// TIA Portal project "EbAndon v2_1_0" (V15) (continued)
   // me.stations[14] : chm 04
   // me.stations[15] : cdo 01
   // me.stations[16] : cdo 02
   // me.stations[17] : cdo 03
   // me.stations[18] : bfl 01
   // me.stations[19] : bfl 02
   // me.stations[20] : bfl 03
   // me.stations[21] : lgs 01
   // me.stations[22] : lgs 02
   // me.stations[23] : lgs 03
   // me.stations[24] : cv 01
   // me.stations[25] : cv 02
   // me.stations[26] : cv 03
   // me.stations[27] : cv 04
   // me.stations[28] : pc 01
   // me.stations[29] : pc 02
END_DATA_BLOCK

// folder: Network Diagnostics

DATA_BLOCK "Net Diag: Global"   // DB7
{ S7_Optimized_Access := 'TRUE' }
VERSION : 0.1
   VAR
      plcData : "UserDiag_typePLC";   // PLC diagnostics data
      ioSystemData : Array[1.."USERDIAG_IO_SYSTEMS_UPPER_LIM"] of "UserDiag_typeIOSystem";   // IO-System diagnostics data
      startDiag : Bool := false;   // Startflag for diagnostic
   END_VAR
BEGIN
END_DATA_BLOCK

DATA_BLOCK "Net Diag: Startup"   // DB8
{ S7_Optimized_Access := 'TRUE' }
VERSION : 0.1
// stored: InstanceOfName NetDiag: Coordinate
"NetDiag: Coordinate"
BEGIN
END_DATA_BLOCK

// folder: (top level)

FUNCTION_BLOCK "EMP"   // FB1, LAD
{ S7_Optimized_Access := 'TRUE' }
VERSION : 0.1
   VAR
      instAniPNTmr : "Animate: PN & Timers";
      instBaseAni : "Base Animations";
      instClrReqData : "Clear Part Requests";
      instClpseTable : "Collapse Table";
      instDfltTmrPrst : "Load Default Timer Presets";
      instHMIAni : "Format Part Call Requests";
      instHMIBarcode : "HMI Barcod Screen";
      instHMISettings : "HMI Settings Screen";
      instInitialize : "Initialize";
      instKP8BtnAct : "KP8 Button Activation";
      instKP8Drvs : Array[0.."stnCount"] of "KP8 Driver";
      instKP8ExpAni : "KP8 Expanded Animations";
      instPartTimers : "Part Timers";
      instPopulateHMI : "HMI Populate Part Call";
      instPopulateLED : "LED Populate Sign";
      instRcrdPartReq : "Record Part Request";
      instRmvPartReq : "Remove Part Request";
      instRstInitReq : "Reset Init Requests";
      instSLAni : "Stack Light Animations";
   END_VAR
   VAR RETAIN
      stations : "Stations";
   END_VAR
   VAR
      instGlblToSim : "Global to Sim";
      instLogReq : "Buffer Log: Part Requests";
      instUserDiag_Diag : "NetDiag: Coordinate";
      instUserDiagGetIPAddress : "NetDiag: Get IPs";
      statStartDiag : Bool := false;   // Static start Diagnostics
      instNetHealthScreen : "HMI: Network Health";
      instHMIStationDriver : "HSS: Driver";
   END_VAR
   VAR_TEMP
      i : Int;
   END_VAR
BEGIN

REGION Network 1: Static start Diagnostics
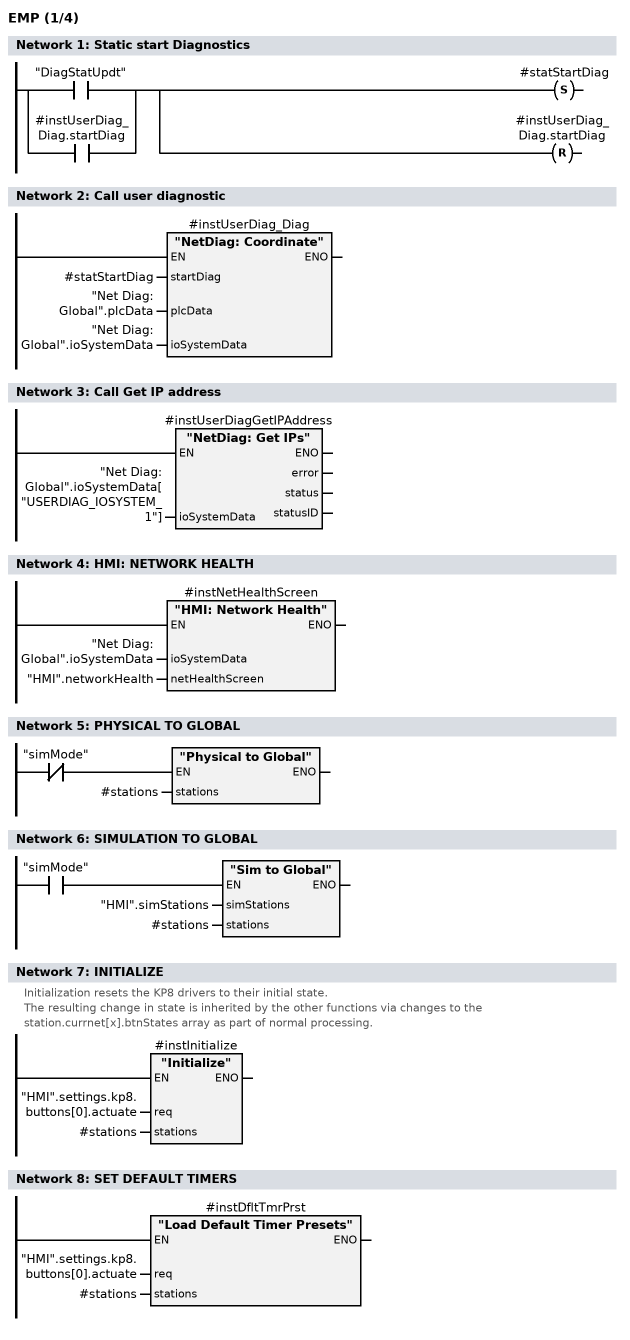
   RUNG wire#powerrail
      Contact( "DiagStatUpdt" )
      wire#w1
      S_Coil( #statStartDiag )
   END_RUNG
   RUNG wire#powerrail
      Contact( #instUserDiag_Diag.startDiag )
   END_RUNG wire#w1
   RUNG wire#w1
      R_Coil( #instUserDiag_Diag.startDiag )
   END_RUNG
   // the same network as SCL:
   IF "DiagStatUpdt" OR #instUserDiag_Diag.startDiag THEN
       #statStartDiag := TRUE;
       #instUserDiag_Diag.startDiag := FALSE;
   END_IF;
END_REGION

REGION Network 2: Call user diagnostic
   RUNG wire#powerrail
      #instUserDiag_Diag(startDiag := #statStartDiag, plcData := "Net Diag: Global".plcData, ioSystemData := "Net Diag: Global".ioSystemData)
   END_RUNG
   // the same network as SCL:
   #instUserDiag_Diag(startDiag := #statStartDiag,   // "NetDiag: Coordinate"
                      plcData := "Net Diag: Global".plcData,
                      ioSystemData := "Net Diag: Global".ioSystemData);
END_REGION

REGION Network 3: Call Get IP address
   RUNG wire#powerrail
      #instUserDiagGetIPAddress(ioSystemData := "Net Diag: Global".ioSystemData["USERDIAG_IOSYSTEM_1"], error =>, status =>, statusID =>)
   END_RUNG
   // the same network as SCL:
   #instUserDiagGetIPAddress(ioSystemData := "Net Diag: Global".ioSystemData["USERDIAG_IOSYSTEM_1"]);   // "NetDiag: Get IPs"
END_REGION

REGION Network 4: HMI: NETWORK HEALTH
   RUNG wire#powerrail
      #instNetHealthScreen(ioSystemData := "Net Diag: Global".ioSystemData, netHealthScreen := "HMI".networkHealth)
   END_RUNG
   // the same network as SCL:
   #instNetHealthScreen(ioSystemData := "Net Diag: Global".ioSystemData, netHealthScreen := "HMI".networkHealth);   // "HMI: Network Health"
END_REGION

REGION Network 5: PHYSICAL TO GLOBAL
   RUNG wire#powerrail
      I_Contact( "simMode" )
      "Physical to Global"(stations := #stations)
   END_RUNG
   // the same network as SCL:
   IF NOT "simMode" THEN "Physical to Global"(stations := #stations); END_IF;
END_REGION

REGION Network 6: SIMULATION TO GLOBAL
   RUNG wire#powerrail
      Contact( "simMode" )
      "Sim to Global"(simStations := "HMI".simStations, stations := #stations)
   END_RUNG
   // the same network as SCL:
   IF "simMode" THEN "Sim to Global"(simStations := "HMI".simStations, stations := #stations); END_IF;
END_REGION

REGION Network 7: INITIALIZE
   // Initialization resets the KP8 drivers to their initial state.
   // The resulting change in state is inherited by the other functions via changes to the
   // station.currnet[x].btnStates array as part of normal processing.
   RUNG wire#powerrail
      #instInitialize(req := "HMI".settings.kp8.buttons[0].actuate, stations := #stations)
   END_RUNG
   // the same network as SCL:
   #instInitialize(req := "HMI".settings.kp8.buttons[0].actuate, stations := #stations);   // "Initialize"
END_REGION

REGION Network 8: SET DEFAULT TIMERS
   RUNG wire#powerrail
      #instDfltTmrPrst(req := "HMI".settings.kp8.buttons[0].actuate, stations := #stations)
   END_RUNG
   // the same network as SCL:
   #instDfltTmrPrst(req := "HMI".settings.kp8.buttons[0].actuate, stations := #stations);   // "Load Default Timer Presets"
END_REGION

REGION Network 9: CLEAR PART REQUEST DATA
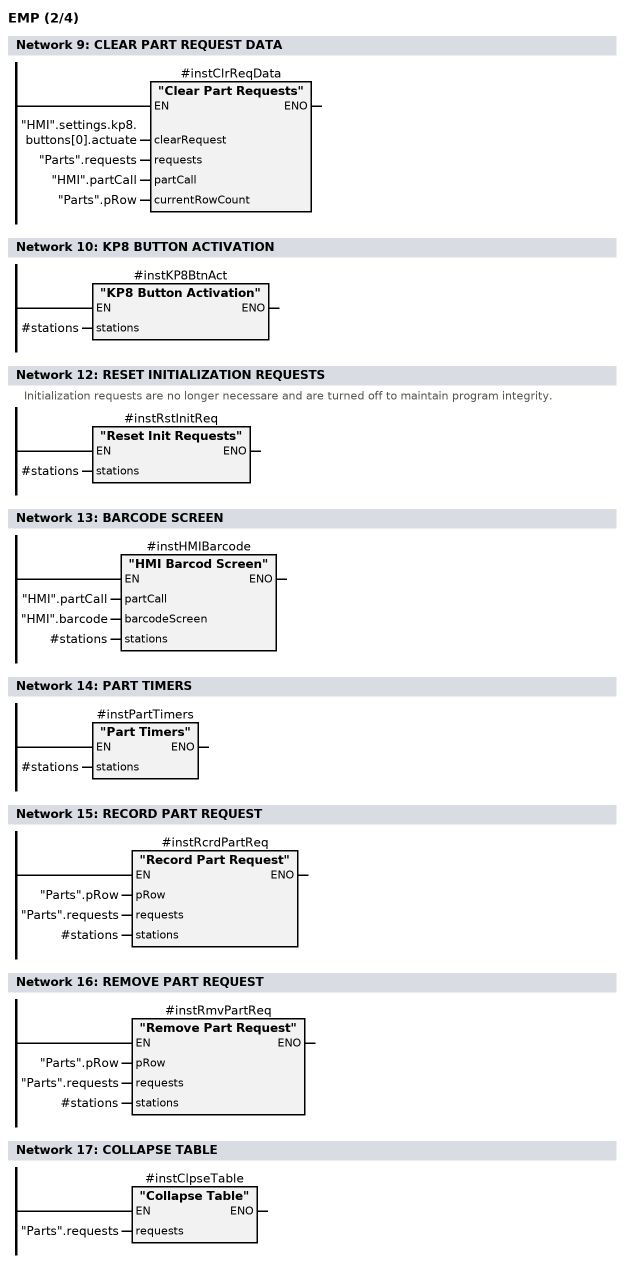
   RUNG wire#powerrail
      #instClrReqData(clearRequest := "HMI".settings.kp8.buttons[0].actuate, requests := "Parts".requests, partCall := "HMI".partCall, currentRowCount := "Parts".pRow)
   END_RUNG
   // the same network as SCL:
   #instClrReqData(clearRequest := "HMI".settings.kp8.buttons[0].actuate,   // "Clear Part Requests"
                   requests := "Parts".requests,
                   partCall := "HMI".partCall,
                   currentRowCount := "Parts".pRow);
END_REGION

REGION Network 10: KP8 BUTTON ACTIVATION
   RUNG wire#powerrail
      #instKP8BtnAct(stations := #stations)
   END_RUNG
   // the same network as SCL:
   #instKP8BtnAct(stations := #stations);   // "KP8 Button Activation"
END_REGION

REGION Network 11 (SCL): KP8 DRIVER CALLS
   REGION "LOOP THROUGH STATIONS"
       FOR #i := 0 TO "stnCount" DO
           #instKP8Drvs[#i](btnIn := #stations.me[#i].kp8In,
                            hardInit := #stations.me[#i].init.hard,
                            softInit := #stations.me[#i].init.soft,
                            btn0Activate := #stations.me[#i].kp8Config.activate[0],
                            btn0Mode := #stations.me[#i].kp8Config.mode[0],
                            btn0Group := #stations.me[#i].kp8Config.group[0],
                            btn0Flash := #stations.me[#i].kp8Config.flash[0],
                            btn0ColorOn1 := #stations.me[#i].kp8Config.colorOn1[0],
                            btn0ColorOn2 := #stations.me[#i].kp8Config.colorOn2[0],
                            btn0ColorOff := #stations.me[#i].kp8Config.colorOff[0],
                            btn1Activate := #stations.me[#i].kp8Config.activate[1],
                            btn1Mode := #stations.me[#i].kp8Config.mode[1],
                            btn1Group := #stations.me[#i].kp8Config.group[1],
                            btn1Flash := #stations.me[#i].kp8Config.flash[1],
                            btn1ColorOn1 := #stations.me[#i].kp8Config.colorOn1[1],
                            btn1ColorOn2 := #stations.me[#i].kp8Config.colorOn2[1],
                            btn1ColorOff := #stations.me[#i].kp8Config.colorOff[1],
                            btn2Activate := #stations.me[#i].kp8Config.activate[2],
                            btn2Mode := #stations.me[#i].kp8Config.mode[2],
                            btn2Group := #stations.me[#i].kp8Config.group[2],
                            btn2Flash := #stations.me[#i].kp8Config.flash[2],
                            btn2ColorOn1 := #stations.me[#i].kp8Config.colorOn1[2],
                            btn2ColorOn2 := #stations.me[#i].kp8Config.colorOn2[2],
                            btn2ColorOff := #stations.me[#i].kp8Config.colorOff[2],
                            btn3Activate := #stations.me[#i].kp8Config.activate[3],
                            btn3Mode := #stations.me[#i].kp8Config.mode[3],
                            btn3Group := #stations.me[#i].kp8Config.group[3],
                            btn3Flash := #stations.me[#i].kp8Config.flash[3],
                            btn3ColorOn1 := #stations.me[#i].kp8Config.colorOn1[3],
                            btn3ColorOn2 := #stations.me[#i].kp8Config.colorOn2[3],
                            btn3ColorOff := #stations.me[#i].kp8Config.colorOff[3],
                            btn4Activate := #stations.me[#i].kp8Config.activate[4],
                            btn4Mode := #stations.me[#i].kp8Config.mode[4],
                            btn4Group := #stations.me[#i].kp8Config.group[4],
                            btn4Flash := #stations.me[#i].kp8Config.flash[4],
                            btn4ColorOn1 := #stations.me[#i].kp8Config.colorOn1[4],
                            btn4ColorOn2 := #stations.me[#i].kp8Config.colorOn2[4],
                            btn4ColorOff := #stations.me[#i].kp8Config.colorOff[4],
                            btn5Activate := #stations.me[#i].kp8Config.activate[5],
                            btn5Mode := #stations.me[#i].kp8Config.mode[5],
                            btn5Group := #stations.me[#i].kp8Config.group[5],
                            btn5Flash := #stations.me[#i].kp8Config.flash[5],
                            btn5ColorOn1 := #stations.me[#i].kp8Config.colorOn1[5],
                            btn5ColorOn2 := #stations.me[#i].kp8Config.colorOn2[5],
                            btn5ColorOff := #stations.me[#i].kp8Config.colorOff[5],
                            btn6Activate := #stations.me[#i].kp8Config.activate[6],
                            btn6Mode := #stations.me[#i].kp8Config.mode[6],
                            btn6Group := #stations.me[#i].kp8Config.group[6],
                            btn6Flash := #stations.me[#i].kp8Config.flash[6],
                            btn6ColorOn1 := #stations.me[#i].kp8Config.colorOn1[6],
                            btn6ColorOn2 := #stations.me[#i].kp8Config.colorOn2[6],
                            btn6ColorOff := #stations.me[#i].kp8Config.colorOff[6],
                            btn7Activate := #stations.me[#i].kp8Config.activate[7],
                            btn7Mode := #stations.me[#i].kp8Config.mode[7],
                            btn7Group := #stations.me[#i].kp8Config.group[7],
                            btn7Flash := #stations.me[#i].kp8Config.flash[7],
                            btn7ColorOn1 := #stations.me[#i].kp8Config.colorOn1[7],
                            btn7ColorOn2 := #stations.me[#i].kp8Config.colorOn2[7],
                            btn7ColorOff := #stations.me[#i].kp8Config.colorOff[7],
                            btnStatesOut => #stations.me[#i].btnStates,
                            btnColorsOut => #stations.me[#i].kp8Out);
       END_FOR;
   END_REGION
END_REGION

REGION Network 12: RESET INITIALIZATION REQUESTS
   // Initialization requests are no longer necessare and are turned off to maintain program integrity.
   RUNG wire#powerrail
      #instRstInitReq(stations := #stations)
   END_RUNG
   // the same network as SCL:
   #instRstInitReq(stations := #stations);   // "Reset Init Requests"
END_REGION

REGION Network 13: BARCODE SCREEN
   RUNG wire#powerrail
      #instHMIBarcode(partCall := "HMI".partCall, barcodeScreen := "HMI".barcode, stations := #stations)
   END_RUNG
   // the same network as SCL:
   #instHMIBarcode(partCall := "HMI".partCall, barcodeScreen := "HMI".barcode, stations := #stations);   // "HMI Barcod Screen"
END_REGION

REGION Network 14: PART TIMERS
   RUNG wire#powerrail
      #instPartTimers(stations := #stations)
   END_RUNG
   // the same network as SCL:
   #instPartTimers(stations := #stations);   // "Part Timers"
END_REGION

REGION Network 15: RECORD PART REQUEST
   RUNG wire#powerrail
      #instRcrdPartReq(pRow := "Parts".pRow, requests := "Parts".requests, stations := #stations)
   END_RUNG
   // the same network as SCL:
   #instRcrdPartReq(pRow := "Parts".pRow, requests := "Parts".requests, stations := #stations);   // "Record Part Request"
END_REGION

REGION Network 16: REMOVE PART REQUEST
   RUNG wire#powerrail
      #instRmvPartReq(pRow := "Parts".pRow, requests := "Parts".requests, stations := #stations)
   END_RUNG
   // the same network as SCL:
   #instRmvPartReq(pRow := "Parts".pRow, requests := "Parts".requests, stations := #stations);   // "Remove Part Request"
END_REGION

REGION Network 17: COLLAPSE TABLE
   RUNG wire#powerrail
      #instClpseTable(requests := "Parts".requests)
   END_RUNG
   // the same network as SCL:
   #instClpseTable(requests := "Parts".requests);   // "Collapse Table"
END_REGION

REGION Network 18: LOG REQUESTS
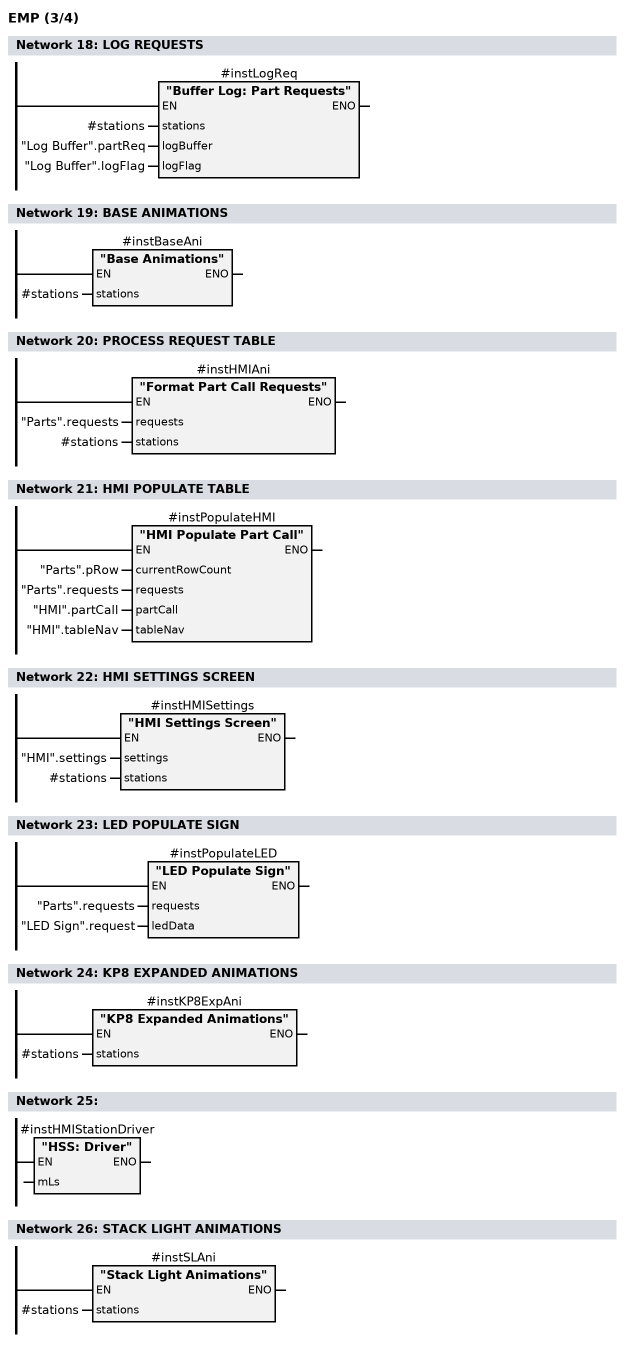
   RUNG wire#powerrail
      #instLogReq(stations := #stations, logBuffer := "Log Buffer".partReq, logFlag := "Log Buffer".logFlag)
   END_RUNG
   // the same network as SCL:
   #instLogReq(stations := #stations, logBuffer := "Log Buffer".partReq, logFlag := "Log Buffer".logFlag);   // "Buffer Log: Part Requests"
END_REGION

REGION Network 19: BASE ANIMATIONS
   RUNG wire#powerrail
      #instBaseAni(stations := #stations)
   END_RUNG
   // the same network as SCL:
   #instBaseAni(stations := #stations);   // "Base Animations"
END_REGION

REGION Network 20: PROCESS REQUEST TABLE
   RUNG wire#powerrail
      #instHMIAni(requests := "Parts".requests, stations := #stations)
   END_RUNG
   // the same network as SCL:
   #instHMIAni(requests := "Parts".requests, stations := #stations);   // "Format Part Call Requests"
END_REGION

REGION Network 21: HMI POPULATE TABLE
   RUNG wire#powerrail
      #instPopulateHMI(currentRowCount := "Parts".pRow, requests := "Parts".requests, partCall := "HMI".partCall, tableNav := "HMI".tableNav)
   END_RUNG
   // the same network as SCL:
   #instPopulateHMI(currentRowCount := "Parts".pRow,   // "HMI Populate Part Call"
                    requests := "Parts".requests,
                    partCall := "HMI".partCall,
                    tableNav := "HMI".tableNav);
END_REGION

REGION Network 22: HMI SETTINGS SCREEN
   RUNG wire#powerrail
      #instHMISettings(settings := "HMI".settings, stations := #stations)
   END_RUNG
   // the same network as SCL:
   #instHMISettings(settings := "HMI".settings, stations := #stations);   // "HMI Settings Screen"
END_REGION

REGION Network 23: LED POPULATE SIGN
   RUNG wire#powerrail
      #instPopulateLED(requests := "Parts".requests, ledData := "LED Sign".request)
   END_RUNG
   // the same network as SCL:
   #instPopulateLED(requests := "Parts".requests, ledData := "LED Sign".request);   // "LED Populate Sign"
END_REGION

REGION Network 24: KP8 EXPANDED ANIMATIONS
   RUNG wire#powerrail
      #instKP8ExpAni(stations := #stations)
   END_RUNG
   // the same network as SCL:
   #instKP8ExpAni(stations := #stations);   // "KP8 Expanded Animations"
END_REGION

REGION Network 25
   RUNG wire#powerrail
      #instHMIStationDriver(mLs :=)
   END_RUNG
   // the same network as SCL:
   #instHMIStationDriver();   // "HSS: Driver"
END_REGION

REGION Network 26: STACK LIGHT ANIMATIONS
   RUNG wire#powerrail
      #instSLAni(stations := #stations)
   END_RUNG
   // the same network as SCL:
   #instSLAni(stations := #stations);   // "Stack Light Animations"
END_REGION

REGION Network 27: GLOBAL TO SIMULATION
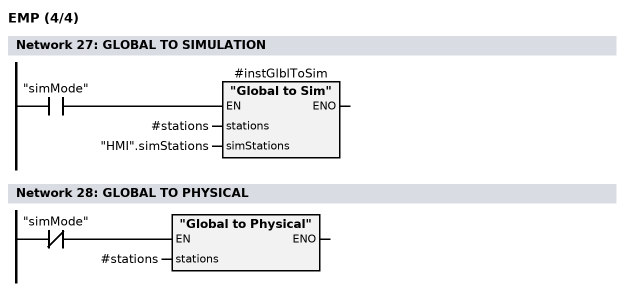
   RUNG wire#powerrail
      Contact( "simMode" )
      #instGlblToSim(stations := #stations, simStations := "HMI".simStations)
   END_RUNG
   // the same network as SCL:
   IF "simMode" THEN
       #instGlblToSim(stations := #stations, simStations := "HMI".simStations);   // "Global to Sim"
   END_IF;
END_REGION

REGION Network 28: GLOBAL TO PHYSICAL
   RUNG wire#powerrail
      I_Contact( "simMode" )
      "Global to Physical"(stations := #stations)
   END_RUNG
   // the same network as SCL:
   IF NOT "simMode" THEN "Global to Physical"(stations := #stations); END_IF;
END_REGION
END_FUNCTION_BLOCK

FUNCTION "Get Recipes Per Station" : Void   // FC30, SCL
{ S7_Optimized_Access := 'TRUE' }
VERSION : 0.1
   VAR_INPUT
      libs : "Menu: Libraries";
   END_VAR
   VAR_TEMP
      i : Int;
      j : Int;
      thisEntry : WString;
      size : Int;
      stn : "Menu: Library";
   END_VAR
   VAR CONSTANT
      blank : WString;
   END_VAR
BEGIN
   FOR #i := 0 TO "stnCount" DO
       #stn := #libs.stations[#i];
       #size := 0;
       FOR #j := 0 TO "menuCntPerStn" DO
           #thisEntry := #stn.entry[#j];
           IF #thisEntry <> #blank THEN
               #size += 1;
           END_IF;
       END_FOR;
       "Recipe Libraries".me.stations[#i].size := #size;
   END_FOR;
END_FUNCTION

// folder: HMI Select Station

FUNCTION_BLOCK "HSS: Driver"   // FB32, LAD
{ S7_Optimized_Access := 'TRUE' }
VERSION : 0.1
   VAR_INPUT
      mLs : "Menu: Libraries";
   END_VAR
   VAR
      recipeSelector : Int;
      r1 : DInt;
      instHSSMenuSelection : "HSS: Menu Selection";
   END_VAR
   VAR_TEMP
      i : Int;
   END_VAR
BEGIN

REGION Network 1
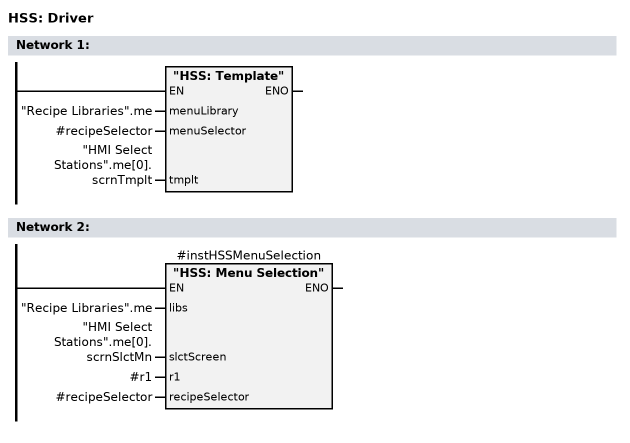
   RUNG wire#powerrail
      "HSS: Template"(menuLibrary := "Recipe Libraries".me, menuSelector := #recipeSelector, tmplt := "HMI Select Stations".me[0].scrnTmplt)
   END_RUNG
   // the same network as SCL:
   "HSS: Template"(menuLibrary := "Recipe Libraries".me,
                   menuSelector := #recipeSelector,
                   tmplt := "HMI Select Stations".me[0].scrnTmplt);
END_REGION

REGION Network 2
   RUNG wire#powerrail
      #instHSSMenuSelection(libs := "Recipe Libraries".me, slctScreen := "HMI Select Stations".me[0].scrnSlctMn, r1 := #r1, recipeSelector := #recipeSelector)
   END_RUNG
   // the same network as SCL:
   #instHSSMenuSelection(libs := "Recipe Libraries".me,   // "HSS: Menu Selection"
                         slctScreen := "HMI Select Stations".me[0].scrnSlctMn,
                         r1 := #r1,
                         recipeSelector := #recipeSelector);
END_REGION
END_FUNCTION_BLOCK

FUNCTION_BLOCK "HSS: Menu Selection"   // FB35, SCL
{ S7_Optimized_Access := 'TRUE' }
VERSION : 0.1
   VAR_INPUT
      libs : "Menu: Libraries";
   END_VAR
   VAR_IN_OUT
      slctScreen : "HSS: Menu Selection Screen";
      r1 : DInt;
      recipeSelector : Int;
   END_VAR
   VAR
      old : Struct
         navPress : Bool;
      END_STRUCT;
      instTableNavigation : "Table Navigatio";
   END_VAR
   VAR_TEMP
      eval : "HSS: Menu Selection Screen";
      pbs : Array[0..#pbFlagCnt] of Bool;
      POS : DInt;
      status : DInt;
      i : Int;
      btnNum : Int;
      pRowVisLbl : Int;
      pRowInvisLbl : Int;
      pRecipeInvisLbl : Int;
      pRecipeVisLbl : Int;
      pRecipeLib : Int;
      pRowTxt : Int;
      pRecipeTxt : Int;
      shifter : DWord;
      btnsAsBool : Array[0..31] of Bool;
      rows : Array[0..99] of DInt;
      offset : DInt;
      navPress : Bool;
      selPress : Bool;
      maxRows : DInt;
   END_VAR
   VAR CONSTANT
      pbFlagCnt : Int := 31;
      btnCnt : Int := 5;
      navMask : DWord := 16#0000_003F;
      visRows : DInt := 6;
      home : DInt := -1000;
      end : DInt := -2000;
   END_VAR
BEGIN
   REGION "INITITALIZE LOCALS"
       #eval := #slctScreen;
       #maxRows := #libs.stations[24].size;
       SCATTER(IN := #eval.pbs,
               OUT => #btnsAsBool);
   END_REGION


   REGION "GET RECIPE SELECTION PRESS" 
       FOR #i := 6 TO 31 DO
           IF #btnsAsBool[#i] THEN
               #recipeSelector := DINT_TO_INT(#r1) + #i - 6;
               #selPress := TRUE;
               EXIT;
           END_IF;
       END_FOR;
   END_REGION


   IF "HMI Select Stations".me[0].scrnSlctMn.pbs.%X0 THEN
       #offset := #home;
   END_IF;
   IF "HMI Select Stations".me[0].scrnSlctMn.pbs.%X1 THEN
       #offset := -1 * #visRows;
   END_IF;
   IF "HMI Select Stations".me[0].scrnSlctMn.pbs.%X2 THEN
       #offset := -1;
   END_IF;
   IF "HMI Select Stations".me[0].scrnSlctMn.pbs.%X3 THEN
       #offset := 1;
   END_IF;
   IF "HMI Select Stations".me[0].scrnSlctMn.pbs.%X4 THEN
       #offset := #visRows;
   END_IF;
   IF "HMI Select Stations".me[0].scrnSlctMn.pbs.%X5 THEN
       #offset := #end;
   END_IF;

   IF ("HMI Select Stations".me[0].scrnSlctMn.pbs AND #navMask) <> 0 THEN
       #navPress := true;
   END_IF;

   REGION "NAV BUTTONS"
       IF #maxRows > #visRows THEN
           FOR #i := 0 TO #btnCnt DO
               #eval.animate[#i] := "BgGray";
               IF #btnsAsBool[#i] THEN
                   #eval.animate[#i] := "BgLTe";
               END_IF;
           END_FOR;
       END_IF;

   END_REGION


   #instTableNavigation(maxRows := #maxRows,
                        visRows := #visRows,
                        offset := #offset,
                        trigger := #navPress,
                        r1 := #r1,
                        rowIndices := #rows);

   IF #navPress AND NOT #old.navPress THEN

       REGION "NARROW ROWS WITH BUTTONS"
           IF #maxRows > #visRows THEN

               REGION "LABELS"
                   FOR #i := 0 TO #visRows - 1 DO

                       #pRowVisLbl := #i + #btnCnt + 1;
                       #pRowInvisLbl := #i + #btnCnt + DINT_TO_INT(#visRows) + 2;
                       #pRecipeLib := #i;
                       #pRowTxt := (#i * 2) + #btnCnt + 1;
                       #pRecipeTxt := #pRowTxt + 1;


                       #eval.animate[#pRowVisLbl] := "BgGray";
                       #eval.animate[#pRowInvisLbl] := "invisible";
                       #eval.txt[#pRowTxt] := "Strip Sign"(DINT_TO_WSTRING(#rows[#i]));
                       #eval.txt[#pRecipeTxt] := "Word Wrap"(stringIn := #libs.stations[24].entry[#rows[#i]],
                                                             maxLength := 22);

                   END_FOR;
               END_REGION

           END_IF;
       END_REGION

       REGION "WIDE ROWS WITHOUT BUTTONS"
           IF #maxRows <= #visRows THEN

               REGION "NAV BUTTONS"
                   FOR #i := 0 TO #btnCnt DO
                       #eval.animate[#i] := "invisible";
                   END_FOR;
               END_REGION

               REGION "LABELS"
                   FOR #i := 0 TO #visRows - 1 DO

                       #pRowVisLbl := #i + #btnCnt + DINT_TO_INT(#visRows) + 2;
                       #pRowInvisLbl := #i + #btnCnt + 1;
                       #pRecipeLib := #i;
                       #pRowTxt := (#i * 2) + #btnCnt + 1;
                       #pRecipeTxt := #pRowTxt + 1;


                       #eval.animate[#pRowVisLbl] := "BgGray";
                       #eval.animate[#pRowInvisLbl] := "invisible";
                       #eval.txt[#pRowTxt] := "Strip Sign"(DINT_TO_WSTRING(#rows[#i]));
                       #eval.txt[#pRecipeTxt] := "Word Wrap"(stringIn := #libs.stations[24].entry[#rows[#i]],
                                                             maxLength := 28);

                   END_FOR;
               END_REGION

           END_IF;
       END_REGION
   END_IF;

   #old.navPress := #navPress;
   #slctScreen := #eval;
END_FUNCTION_BLOCK

FUNCTION "HSS: Template" : Void   // FC24, SCL
{ S7_Optimized_Access := 'TRUE' }
VERSION : 0.1
   VAR_INPUT
      menuLibrary : "Menu: Libraries";
      menuSelector : Int;
   END_VAR
   VAR_IN_OUT
      tmplt : "HSS: Template Screen";
   END_VAR
   VAR_TEMP
      i : Int;
   END_VAR
BEGIN
   #tmplt.animate[0] := "BgGray";
   #tmplt.text[0] := "Word Wrap"(stringIn := #menuLibrary.stations[24].entry[#menuSelector],
                                 maxLength := 26);
END_FUNCTION

// folder: Network Diagnostics

FUNCTION_BLOCK "NetDiag: Get IPs"   // FB27, SCL
{ S7_Optimized_Access := 'TRUE' }
VERSION : 0.1
   VAR_OUTPUT
      error : Bool := FALSE;   // Rising edge informs that an error occurred during the execution of the FB
      status : Word := 16#0000;   // Current status of FB
      statusID : Word := 16#0;   // Current status ID of calling instruction
   END_VAR
   VAR_IN_OUT
      ioSystemData : "UserDiag_typeIOSystem";   // IO-System diagnostics data
   END_VAR
   VAR
      statError : Bool := FALSE;   // Static value for output error
      statStatus : Word := 16#0000;   // Static value for output status
      statStatusID : Word := 16#0;   // Static value for output statusID
      instGetStationInfo : GetStationInfo;   // Instance of GetStationInfo
      statFirstDeviceFlag : Bool := TRUE;   // Help tag for the first device in the linked list
      statDeviceIndex : Int := 0;   // Device/slave index
   END_VAR
   VAR_TEMP
      tempIP : IF_CONF_v4;   // Temporary IP address
   END_VAR
   VAR CONSTANT
      STATUS_EXECUTION_FINISHED : Word := 16#0000;   // Execution finished without errors
      ID_GET_STATION_INFO : Word := 12;   // StatusID during GetStationInfo command
      MODE_IPV4 : UInt := 1;   // Address parameter according to IPv4
      LAST_DEVICE : Int := -1;   // No next device
   END_VAR
BEGIN
   //=============================================================================
   //SIEMENS AG
   //(c)Copyright 2015 All Rights Reserved
   //-----------------------------------------------------------------------------
   //Library: 
   //Tested with: S7-1516-3 PN/DP FW 2.5
   //Engineering: TIA Portal V15
   //Restrictions: Call in cyclic OB
   //Requirements: -
   //Functionality: Get IP address of IO devices
   //-----------------------------------------------------------------------------
   //Change log table:
   //Version  Date       Expert in charge                Changes applied
   //01.00.00 20.12.2017 Siemens Industry Online Support First released version
   //=============================================================================

   //=============================================================================
   // Go through existing devices and get IP address
   //=============================================================================
   // Initialize the pointer for the first run 
   IF (#statFirstDeviceFlag = TRUE)
   THEN
       #statDeviceIndex := #ioSystemData.firstDevice;
       #statFirstDeviceFlag := FALSE;
   END_IF;

   // Check and store the IP address, if the device is existing
   // GetStationInfo is an acyclic instruction. In the FB, the
   // instruction has to be repeated until it is done or error
   IF ((#ioSystemData.number >= 100)
       AND (#ioSystemData.number <= 115)
       AND (#ioSystemData.devices[#statDeviceIndex].exists = TRUE)
       AND (#ioSystemData.devices[#statDeviceIndex].ipAddress.ADDR[1] = 0))
   THEN
       // Get IP address of each decive in PN System
       #instGetStationInfo(REQ := TRUE,
                           LADDR := #ioSystemData.devices[#statDeviceIndex].hardwareId,
                           MODE := #MODE_IPV4,
                           DATA := #tempIP);

       IF (#instGetStationInfo.ERROR = TRUE)
       THEN
           // Error handling
           #statStatus := #instGetStationInfo.STATUS;
           #statStatusID := #ID_GET_STATION_INFO;
           #statError := TRUE;

           // Everything is ok --> Copy IP address    
       ELSIF (#instGetStationInfo.DONE = TRUE)
       THEN
           #ioSystemData.devices[#statDeviceIndex].ipAddress := #tempIP.InterfaceAddress;

           // Initialize the pointer for the next run
           #statDeviceIndex := #ioSystemData.devices[#statDeviceIndex].nextDevice;
       ELSE
           ;
       END_IF;
   ELSE
       // Initialize the pointer for the next run
       #statDeviceIndex := #ioSystemData.devices[#statDeviceIndex].nextDevice;
   END_IF;

   // Check last device
   IF (#statDeviceIndex = #LAST_DEVICE)
   THEN
       #statDeviceIndex := #ioSystemData.firstDevice;
   END_IF;

   // Write static values to outputs
   #error := #statError;
   #status := #statStatus;
   #statusID := #statStatusID;
END_FUNCTION_BLOCK

